// ===== library: CodeBlockByCopyVersionObject "None" =====

// ===== library: CodeBlockByCopyVersionObject "None" =====

// ===== library: CodeBlockByCopyVersionObject "None" =====

(* ===== HMI "HMI_RT_1" =====
system functions are stored by id; their names below are inferred from use
connection "HMI_Collegamento_1": ETHERNET, S7_1500_OMS

HMI tags "Tabella delle variabili standard"
   "DB_AUX_AXIS1" : IAI_PCONPRT = PLC DB_AUX.AXIS1, 100 ms
   "DB_AUX_TARGET_POS" : Array [0..4] of DInt = PLC DB_AUX.TARGET_POS AT %DB1.DBW0, 100 ms
   "DB_AUX_HMI_Bit_HMIb1" : Bool = PLC DB_AUX.HMI_Bit.HMIb1 AT %DB1.DBW0, 100 ms
   "DB_AUX_HMI_Bit_HMIb2" : Bool = PLC DB_AUX.HMI_Bit.HMIb2 AT %DB1.DBW0, 100 ms
   "DB_AUX_HMI_Bit_HMIb3" : Bool = PLC DB_AUX.HMI_Bit.HMIb3 AT %DB1.DBW0, 100 ms
   "DB_AUX_HMI_Bit_HMIb4" : Bool = PLC DB_AUX.HMI_Bit.HMIb4 AT %DB1.DBW0, 100 ms
   "DB_AUX_HMI_Bit_HMIb5" : Bool = PLC DB_AUX.HMI_Bit.HMIb5 AT %DB1.DBW0, 100 ms
   "DB_AUX_HMI_Bit_HMIb6" : Bool = PLC DB_AUX.HMI_Bit.HMIb6 AT %DB1.DBW0, 100 ms
   "DB_AUX_HMI_Bit_HMIb7" : Bool = PLC DB_AUX.HMI_Bit.HMIb7 AT %DB1.DBW0, 100 ms
   "DB_AUX_HMI_Bit_HMIb8" : Bool = PLC DB_AUX.HMI_Bit.HMIb8 AT %DB1.DBW0, 100 ms
   "DB_AUX_HMI_Bit_HMIb9" : Bool = PLC DB_AUX.HMI_Bit.HMIb9 AT %DB1.DBW0, 100 ms
   "DB_AUX_HMI_Bit_HMIb10" : Bool = PLC DB_AUX.HMI_Bit.HMIb10 AT %DB1.DBW0, 100 ms
   "DB_AUX_HMI_Bit_HMIb11" : Bool = PLC DB_AUX.HMI_Bit.HMIb11 AT %DB1.DBW0, 100 ms
   "DB_AUX_HMI_Bit_HMIb12" : Bool = PLC DB_AUX.HMI_Bit.HMIb12 AT %DB1.DBW0, 100 ms
   "DB_AUX_HMI_Bit_HMIb13" : Bool = PLC DB_AUX.HMI_Bit.HMIb13 AT %DB1.DBW0, 100 ms
   "DB_AUX_SPEED_POS" : Array [0..4] of UDInt = PLC DB_AUX.SPEED_POS AT %DB1.DBW0, 100 ms
   "DB_AUX_ACC_DEC" : USInt = PLC DB_AUX.ACC_DEC AT %DB1.DBW0, 100 ms

screen "Pagina_1" 800x480
   IOField "Campo I/O_3" at 8,24 size 129x52; FormatPattern s999999
      ProcessValue <- "[1]"
   TextField "Casella di testo_3" at 0,0 size 148x23; Text 'STARTING POS.'
   IOField "Campo I/O_9" at 8,432 size 145x44; FormatPattern 999999
      ProcessValue <- "Current_POS"
   TextField "Casella di testo_11" at 0,408 size 87x23; Text 'POS. FBK'
   IOField "Campo I/O_10" at 160,432 size 97x44; FormatPattern FFFF
      ProcessValue <- "Alarm_COD"
   TextField "Casella di testo_12" at 152,408 size 97x23; Text 'ERR CODE'
   GraphicIOField "PlotLight_Round_R" at 256,432 size 42x42; PictureOn "PilotLight_Round_R_On_256c"; PictureOff "PilotLight_Round_GN_Off_256c"
      ProcessValue <- "CTRL2_Sig_ALM"
   GraphicIOField "PlotLight_Round_R_1" at 558,432 size 42x42; PictureOff "PilotLight_Round_GN_Off_256c"; PictureOn "PilotLight_Round_R_On_256c"
      ProcessValue <- "CTRL2_Sig_MOVE"
   TextField "Casella di testo_13" at 504,408 size 148x23; Text 'AXS IN MOTION'
   TextField "Casella di testo_14" at 648,408 size 152x23; Text 'PROCESS COMP.'
   TextField "Casella di testo_15" at 0,208 size 97x23; Text 'SERVO ON'
   Button "Pulsante_1" at 8,232 size 128x48; TextOff 'ENABLE'
      on Press: InvertBit("DB_AUX_HMI_Bit_HMIb5")
   TextField "Casella di testo_16" at 152,208 size 134x23; Text 'START POSIT.'
   Button "Pulsante_2" at 160,232 size 128x48; TextOff 'START'
      on Press: SetBit("DB_AUX_HMI_Bit_HMIb6")
      on Release: ResetBit("DB_AUX_HMI_Bit_HMIb6")
   TextField "Casella di testo_18" at 16,304 size 86x23; Text 'JOG FWD'
   Button "Pulsante_4" at 8,328 size 104x40; TextOff 'JOG FWD'
      on Press: SetBit("DB_AUX_HMI_Bit_HMIb8")
      on Release: ResetBit("DB_AUX_HMI_Bit_HMIb8")
   TextField "Casella di testo_19" at 128,304 size 82x23; Text 'JOG REV'
   Button "Pulsante_5" at 120,328 size 104x40; TextOff 'JOG REV'
      on Press: SetBit("DB_AUX_HMI_Bit_HMIb9")
      on Release: ResetBit("DB_AUX_HMI_Bit_HMIb9")
   Button "Pulsante_7" at 400,200 size 104x80; TextOff 'HOME'
      on Press: SetBit("DB_AUX_HMI_Bit_HMIb7")
      on Release: ResetBit("DB_AUX_HMI_Bit_HMIb7")
   TextField "Casella di testo_21" at 392,176 size 124x23; Text 'HOME START'
   IOField "Campo I/O_12" at 160,24 size 129x52; FormatPattern s999999
      ProcessValue <- "[2]"
   TextField "Casella di testo_1" at 152,0 size 131x23; Text 'PICKING POS.'
   IOField "Campo I/O_13" at 312,24 size 129x52; FormatPattern s999999
      ProcessValue <- "[3]"
   TextField "Casella di testo_2" at 304,0 size 147x23; Text 'OUT JAWS POS.'
   IOField "Campo I/O_14" at 464,24 size 129x52; FormatPattern s999999
      ProcessValue <- "[4]"
   TextField "Casella di testo_9" at 456,0 size 141x23; Text 'APPROCH.POS.'
   TextField "Casella di testo_4" at 592,0 size 168x23; Text 'LOAD POS->PCON'
   Button "Pulsante_3" at 600,24 size 96x48; TextOff 'STARTING'
      on Press: SetBit("DB_AUX_HMI_Bit_HMIb1")
      on Release: ResetBit("DB_AUX_HMI_Bit_HMIb1")
   Button "Pulsante_8" at 696,24 size 96x48; TextOff 'PICKING'
      on Press: SetBit("DB_AUX_HMI_Bit_HMIb2")
      on Release: ResetBit("DB_AUX_HMI_Bit_HMIb2")
   Button "Pulsante_9" at 600,72 size 96x48; TextOff 'OUT JAWS'
      on Press: SetBit("DB_AUX_HMI_Bit_HMIb3")
      on Release: ResetBit("DB_AUX_HMI_Bit_HMIb3")
   Button "Pulsante_10" at 696,72 size 96x48; TextOff 'APPROCH'
      on Press: SetBit("DB_AUX_HMI_Bit_HMIb4")
      on Release: ResetBit("DB_AUX_HMI_Bit_HMIb4")
   IOField "Campo I/O_1" at 696,120 size 97x36; FormatPattern s999999
      ProcessValue <- "Target_POS"
   TextField "Casella di testo_5" at 8,80 size 92x23; Text 'SPEED P1'
   IOField "Campo I/O_2" at 8,104 size 129x36; FormatPattern 999999
      ProcessValue <- "[1]"
   TextField "Casella di testo_6" at 160,80 size 92x23; Text 'SPEED P2'
   IOField "Campo I/O_4" at 160,104 size 129x36; FormatPattern 999999
      ProcessValue <- "[2]"
   TextField "Casella di testo_7" at 312,80 size 92x23; Text 'SPEED P3'
   IOField "Campo I/O_5" at 312,104 size 129x36; FormatPattern 999999
      ProcessValue <- "[3]"
   TextField "Casella di testo_8" at 464,80 size 92x23; Text 'SPEED P4'
   IOField "Campo I/O_6" at 464,104 size 129x36; FormatPattern 999999
      ProcessValue <- "[4]"
   TextField "Casella di testo_10" at 600,128 size 82x23; Text 'TARG.POS'
   IOField "Campo I/O_7" at 696,152 size 97x36; FormatPattern 999999
      ProcessValue <- "Positioning_BAND"
   TextField "Casella di testo_17" at 600,160 size 87x23; Text 'POS. BAND'
   IOField "Campo I/O_8" at 696,184 size 97x36; FormatPattern 999999
      ProcessValue <- "Speed"
   TextField "Casella di testo_22" at 600,192 size 52x23; Text 'SPEED'
   TextField "Casella di testo_23" at 8,144 size 88x23; Text 'ACC/DEC'
   IOField "Campo I/O_11" at 8,168 size 129x36; FormatPattern 99
      ProcessValue <- "DB_AUX_ACC_DEC"
   TextField "Casella di testo_24" at 600,224 size 72x23; Text 'ACC/DEC'
   IOField "Campo I/O_15" at 696,216 size 97x36; FormatPattern 9999
      ProcessValue <- "Acceleration"
   GraphicIOField "PlotLight_Round_R_2" at 536,216 size 42x42; PictureOff "PilotLight_Round_GN_Off_256c"; PictureOn "PilotLight_Round_GN_On_256c"
      ProcessValue <- "CTRL2_Sig_HEND"
   TextField "Casella di testo_20" at 512,176 size 88x23; Text 'HOME OK'
   GraphicIOField "PlotLight_Round_R_3" at 704,432 size 42x42; PictureOn "PilotLight_Round_GN_On_256c"; PictureOff "PilotLight_Round_GN_Off_256c"
      ProcessValue <- "CTRL2_Sig_PEND"
   Button "Pulsante_6" at 304,432 size 72x48; TextOff 'RES'
      on Release: ResetBit("DB_AUX_HMI_Bit_HMIb10")
      on Press: SetBit("DB_AUX_HMI_Bit_HMIb10")
   TextField "Casella di testo_25" at 296,408 size 84x23; Text 'RES.ALM'
*)